// TIA Portal project "ProjektSklepu" (V18)

(* hardware
DEVICE "S7-1200 station_1"  S7-1200 Station
   slot 0: "Rack_0"  S7-1200 Rack  Rack  V1.0
   slot 1: "PLC_1"  CPU 1214C AC/DC/Rly  6ES7 214-1BG40-0XB0  V4.6
DEVICE "HMI_1"  KTP700 Basic PN
   slot 0: "HMI_1"  KTP700 Basic PN  6AV2 123-2GB03-0AX0  17.0.0.0
   slot 1: "HMI_RT_1"  KTP700 Basic PN  6AV2 123-2GB03-0AX0  17.0.0.0
   slot 5: "HMI_1.IE_CP_1"  PROFINET Interface  17.0.0.0
      slot 1: "PROFINET Interface_1"  PROFINET Interface
         slot 1: "Port_1"  Port
*)

// ===== PLC "PLC_1"  CPU 1214C AC/DC/Rly =====

VAR_GLOBAL   // PLC tag table "TT_Drzwi"
   "CzujnikRuchu_DrzwiWejscie" AT %M0.0 : Bool;
   "SygnalPracownikaDoOtwarcia_DrzwiWejscie" AT %M0.1 : Bool;
   "ZmiennaDoSymulacjiCzujnikaRuchu" AT %M0.2 : Bool;
   "StanDrzwi" AT %M0.7 : Bool;
   "Clock_Byte" AT %MB100 : Byte;
   "Clock_10Hz" AT %M100.0 : Bool;
   "Clock_5Hz" AT %M100.1 : Bool;
   "Clock_2.5Hz" AT %M100.2 : Bool;
   "Clock_2Hz" AT %M100.3 : Bool;
   "Clock_1.25Hz" AT %M100.4 : Bool;
   "Clock_1Hz" AT %M100.5 : Bool;
   "Clock_0.625Hz" AT %M100.6 : Bool;
   "Clock_0.5Hz" AT %M100.7 : Bool;
   "CzujnikRuchuWyjscie" AT %M101.0 : Bool;
   "SygnalPracownikaDoWyjscie" AT %M101.1 : Bool;
   "Liczba osob" AT %MW6 : Int;
   "zmienna pomocnicza do wentylacji" AT %M8.1 : Bool;
   "ZmiennaPomocnicza do zliczania osob" AT %M8.2 : Bool;
   "ZmiennaPomocnicza do zliczania osob wyjscie" AT %M8.3 : Bool;
   "Odliczanie" AT %M8.4 : Bool;
   "StanDrzwiINT" AT %MW4 : Int;
END_VAR

VAR_GLOBAL   // PLC tag table "TT_Temperatura"
   "Grzanie" AT %M0.3 : Bool;
   "Chłodzenie" AT %M0.4 : Bool;
   "ZmiennaPomocnicznaDoGrzania" AT %M0.5 : Bool;
   "ZmiennaPomocniczaDoChłodzenia" AT %M0.6 : Bool;
END_VAR

VAR_GLOBAL   // PLC tag table "TT_Pozar"
   "Tlo" AT %M1.0 : Bool;
   "PrzyciskDoSymulacjiCzujnikaDymu" AT %M1.1 : Bool;
   "CzujnikDymu" AT %M1.2 : Bool;
   "Swiatlo alarmowe" AT %M1.3 : Bool;
   "PracownikAlarm" AT %M1.4 : Bool;
   "ALARM" AT %M1.5 : Bool;
   "Zmienna pomocnicza do swiatla alarmu" AT %M1.6 : Bool;
   "ZmiennaDoSymulacjiCzujnikaWyjscie" AT %M1.7 : Bool;
   "Wlacz wentylacje" AT %M2.0 : Bool;
END_VAR

DATA_BLOCK "Przycisk_DB"   // DB1
{ S7_Optimized_Access := 'TRUE' }
VERSION : 0.1
// stored: InstanceOfName Przycisk
"Przycisk"
BEGIN
END_DATA_BLOCK

DATA_BLOCK "Temperatura"   // DB4
{ S7_Optimized_Access := 'TRUE' }
VERSION : 0.1
   VAR
      TemperaturaAktualna : Int := 15;
      TemperaturaDanaPrzezPracownika : Int := 15;
   END_VAR
BEGIN
END_DATA_BLOCK

DATA_BLOCK "Przycisk_DB_1"   // DB5
{ S7_Optimized_Access := 'TRUE' }
VERSION : 0.1
// stored: InstanceOfName Przycisk
"Przycisk"
BEGIN
END_DATA_BLOCK

DATA_BLOCK "Przycisk_DB_2"   // DB6
{ S7_Optimized_Access := 'TRUE' }
VERSION : 0.1
// stored: InstanceOfName Przycisk
"Przycisk"
BEGIN
END_DATA_BLOCK

DATA_BLOCK "Block_1_DB"   // DB7
{ S7_Optimized_Access := 'TRUE' }
VERSION : 0.1
// stored: InstanceOfName ZmianaBoolNaInt
"ZmianaBoolNaInt"
BEGIN
END_DATA_BLOCK

DATA_BLOCK "Przycisk_DB_3"   // DB8
{ S7_Optimized_Access := 'TRUE' }
VERSION : 0.1
// stored: InstanceOfName Przycisk
"Przycisk"
BEGIN
END_DATA_BLOCK

DATA_BLOCK "Block_1_DB_1"   // DB9
{ S7_Optimized_Access := 'TRUE' }
VERSION : 0.1
// stored: InstanceOfName ZmianaBoolNaInt
"ZmianaBoolNaInt"
BEGIN
END_DATA_BLOCK

// folder: System blocks/Program resources

DATA_BLOCK "IEC_Timer_0_DB"   // DB2
{ S7_Optimized_Access := 'TRUE' }
AUTHOR : Simatic
FAMILY : IEC
NAME : IEC_TMR
VERSION : 1.0
// stored: InstanceOfName IEC_TIMER
"IEC_TIMER"
BEGIN
END_DATA_BLOCK

DATA_BLOCK "IEC_Timer_0_DB_1"   // DB3
{ S7_Optimized_Access := 'TRUE' }
AUTHOR : Simatic
FAMILY : IEC
NAME : IEC_TMR
VERSION : 1.0
// stored: InstanceOfName IEC_TIMER
"IEC_TIMER"
BEGIN
END_DATA_BLOCK

DATA_BLOCK "IEC_Timer_0_DB_4"   // DB10
{ S7_Optimized_Access := 'TRUE' }
AUTHOR : Simatic
FAMILY : IEC
NAME : IEC_TMR
VERSION : 1.0
// stored: InstanceOfName IEC_TIMER
"IEC_TIMER"
BEGIN
END_DATA_BLOCK

// folder: (top level)

FUNCTION_BLOCK "Przycisk"   // FB1, SCL
{ S7_Optimized_Access := 'TRUE' }
VERSION : 0.1
   VAR_INPUT
      HMI_Przycisk : Bool;
   END_VAR
   VAR_IN_OUT
      Lampka : Bool;
   END_VAR
   VAR
      Prev_HMI_Button : Bool;
   END_VAR
BEGIN
   IF #HMI_Przycisk AND NOT #Prev_HMI_Button THEN
       #Lampka := NOT #Lampka;
   END_IF;

   #Prev_HMI_Button := #HMI_Przycisk;
END_FUNCTION_BLOCK

FUNCTION_BLOCK "ZmianaBoolNaInt"   // FB2, SCL
{ S7_Optimized_Access := 'TRUE' }
VERSION : 0.1
   VAR_INPUT
      StanDrzwi : Bool;
   END_VAR
   VAR_OUTPUT
      StanDrzwiInt : Int;
   END_VAR
BEGIN
   IF "StanDrzwi" THEN
       #StanDrzwiInt := 1;
   ELSE
       #StanDrzwiInt := 0;
   END_IF;
END_FUNCTION_BLOCK

ORGANIZATION_BLOCK "Main"   // OB1, LAD, ProgramCycle
TITLE = "Main Program Sweep (Cycle)"
{ S7_Optimized_Access := 'TRUE' }
VERSION : 0.1
   VAR_INPUT
      Initial_Call : Bool;   // Initial call of this OB
      Remanence : Bool;   // =True, if remanent data are available
   END_VAR
   VAR_TEMP   // added for the SCL form of the ladder/FBD networks
      _w1 : Bool;
      _w2 : Bool;
   END_VAR
BEGIN

REGION Network 1: Zmienia stan czujnika wejścia za każdym razem, gdy przycisk zostanie naciśnięty - na zbocze narastające
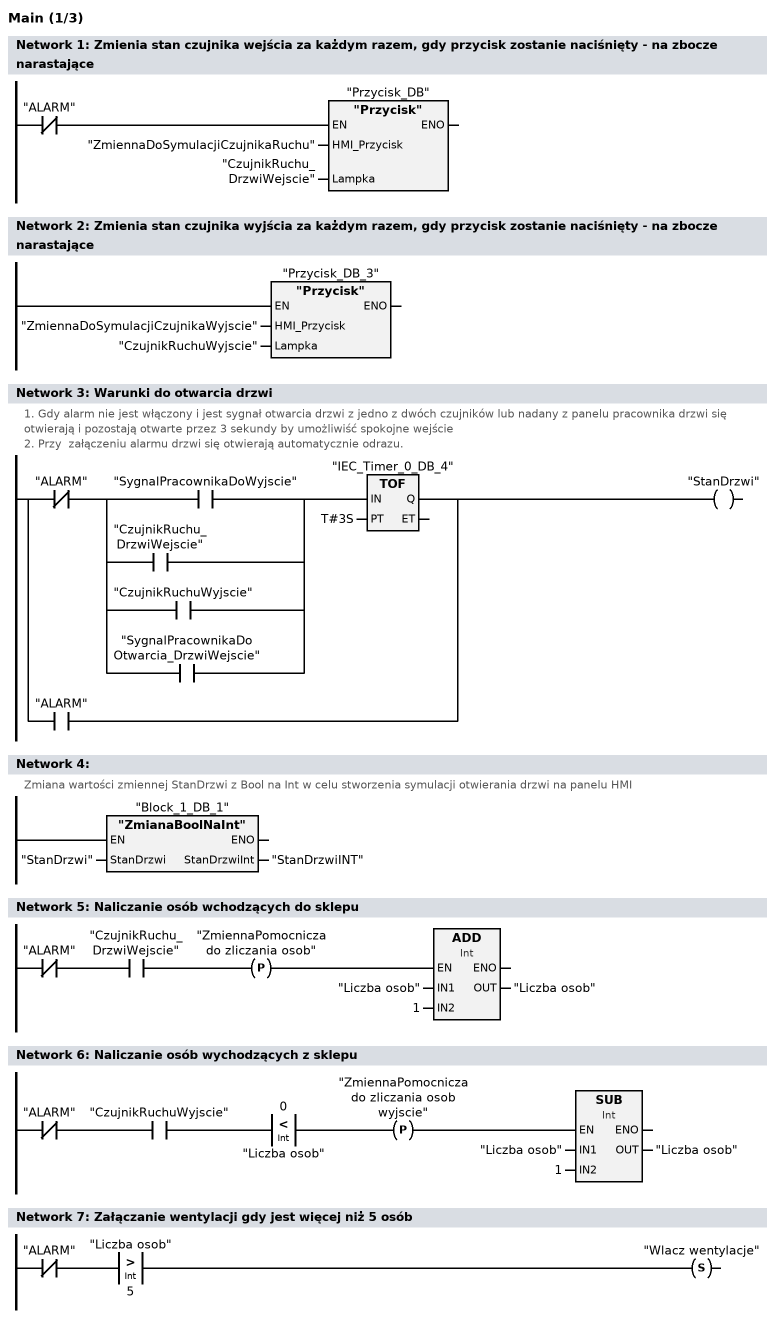
   RUNG wire#powerrail
      I_Contact( "ALARM" )
      "Przycisk_DB"(HMI_Przycisk := "ZmiennaDoSymulacjiCzujnikaRuchu", Lampka := "CzujnikRuchu_DrzwiWejscie")
   END_RUNG
   // the same network as SCL:
   IF NOT "ALARM" THEN
       "Przycisk_DB"(HMI_Przycisk := "ZmiennaDoSymulacjiCzujnikaRuchu", Lampka := "CzujnikRuchu_DrzwiWejscie");   // "Przycisk"
   END_IF;
END_REGION

REGION Network 2: Zmienia stan czujnika wyjścia za każdym razem, gdy przycisk zostanie naciśnięty - na zbocze narastające
   RUNG wire#powerrail
      "Przycisk_DB_3"(HMI_Przycisk := "ZmiennaDoSymulacjiCzujnikaWyjscie", Lampka := "CzujnikRuchuWyjscie")
   END_RUNG
   // the same network as SCL:
   "Przycisk_DB_3"(HMI_Przycisk := "ZmiennaDoSymulacjiCzujnikaWyjscie", Lampka := "CzujnikRuchuWyjscie");   // "Przycisk"
END_REGION

REGION Network 3: Warunki do otwarcia drzwi
   // 1. Gdy alarm nie jest włączony i jest sygnał otwarcia drzwi z jedno z dwóch czujników lub nadany z panelu pracownika drzwi się otwierają i pozostają otwarte przez 3 sekundy by umożliwiść spokojne wejście
   // 2. Przy  załączeniu alarmu drzwi się otwierają automatycznie odrazu.
   "IEC_Timer_0_DB_4".TOF(IN := NOT "ALARM" AND ("SygnalPracownikaDoWyjscie" OR "CzujnikRuchu_DrzwiWejscie" OR "CzujnikRuchuWyjscie" OR "SygnalPracownikaDoOtwarcia_DrzwiWejscie"),
                          PT := T#3S);
   "StanDrzwi" := "IEC_Timer_0_DB_4".Q OR "ALARM";
END_REGION

REGION Network 4
   // Zmiana wartości zmiennej StanDrzwi z Bool na Int w celu stworzenia symulacji otwierania drzwi na panelu HMI
   RUNG wire#powerrail
      "Block_1_DB_1"(StanDrzwi := "StanDrzwi", StanDrzwiInt => "StanDrzwiINT")
   END_RUNG
   // the same network as SCL:
   "Block_1_DB_1"(StanDrzwi := "StanDrzwi", StanDrzwiInt => "StanDrzwiINT");   // "ZmianaBoolNaInt"
END_REGION

REGION Network 5: Naliczanie osób wchodzących do sklepu
   RUNG wire#powerrail
      I_Contact( "ALARM" )
      Contact( "CzujnikRuchu_DrzwiWejscie" )
      P_Trig( "ZmiennaPomocnicza do zliczania osob" )
      { S7_Templates := "SrcType := Int" } Add(in1 := "Liczba osob", in2 := 1, out => "Liczba osob")
   END_RUNG
   // the same network as SCL:
   #_w1 := NOT "ALARM" AND "CzujnikRuchu_DrzwiWejscie";
   #_w2 := #_w1 AND NOT "ZmiennaPomocnicza do zliczania osob";   // rising edge
   "ZmiennaPomocnicza do zliczania osob" := #_w1;
   IF #_w2 THEN "Liczba osob" := "Liczba osob" + 1; END_IF;
END_REGION

REGION Network 6: Naliczanie osób wychodzących z sklepu
   RUNG wire#powerrail
      I_Contact( "ALARM" )
      Contact( "CzujnikRuchuWyjscie" )
      { S7_Templates := "SrcType := Int" } LT_Contact(in1 := 0, in2 := "Liczba osob")
      P_Trig( "ZmiennaPomocnicza do zliczania osob wyjscie" )
      { S7_Templates := "SrcType := Int" } Sub(in1 := "Liczba osob", in2 := 1, out => "Liczba osob")
   END_RUNG
   // the same network as SCL:
   #_w1 := NOT "ALARM" AND "CzujnikRuchuWyjscie" AND (0 < "Liczba osob");
   #_w2 := #_w1 AND NOT "ZmiennaPomocnicza do zliczania osob wyjscie";   // rising edge
   "ZmiennaPomocnicza do zliczania osob wyjscie" := #_w1;
   IF #_w2 THEN "Liczba osob" := "Liczba osob" - 1; END_IF;
END_REGION

REGION Network 7: Załączanie wentylacji gdy jest więcej niż 5 osób
   RUNG wire#powerrail
      I_Contact( "ALARM" )
      { S7_Templates := "SrcType := Int" } GT_Contact(in1 := "Liczba osob", in2 := 5)
      S_Coil( "Wlacz wentylacje" )
   END_RUNG
   // the same network as SCL:
   IF NOT "ALARM" AND ("Liczba osob" > 5) THEN "Wlacz wentylacje" := TRUE; END_IF;
END_REGION

REGION Network 8: Wyłączanie wentylacji gdy jest mniej niz 5 osób
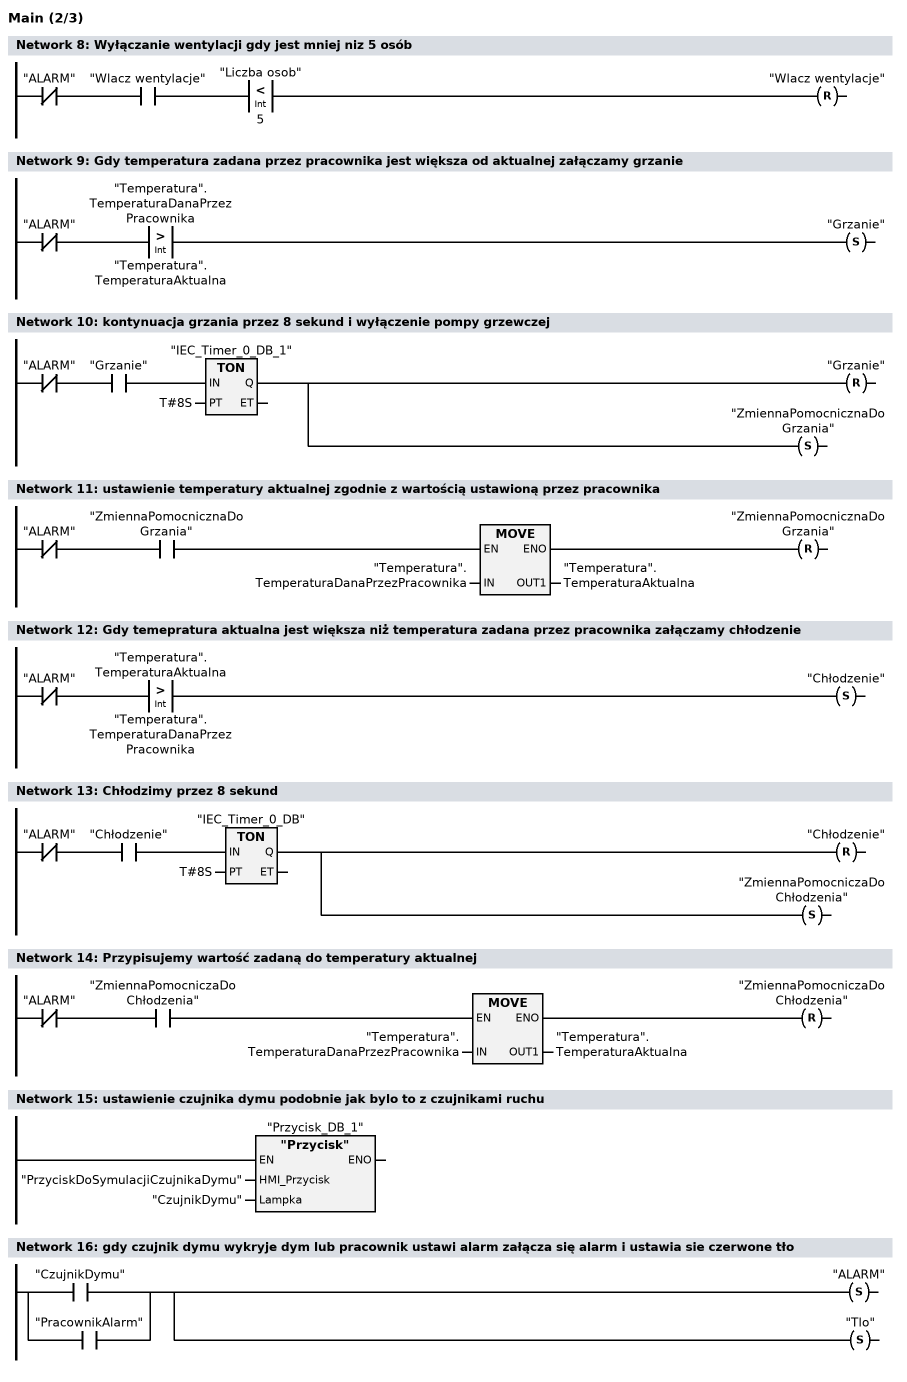
   RUNG wire#powerrail
      I_Contact( "ALARM" )
      Contact( "Wlacz wentylacje" )
      { S7_Templates := "SrcType := Int" } LT_Contact(in1 := "Liczba osob", in2 := 5)
      R_Coil( "Wlacz wentylacje" )
   END_RUNG
   // the same network as SCL:
   IF NOT "ALARM" AND "Wlacz wentylacje" AND ("Liczba osob" < 5) THEN "Wlacz wentylacje" := FALSE; END_IF;
END_REGION

REGION Network 9: Gdy temperatura zadana przez pracownika jest większa od aktualnej załączamy grzanie
   RUNG wire#powerrail
      I_Contact( "ALARM" )
      { S7_Templates := "SrcType := Int" } GT_Contact(in1 := "Temperatura".TemperaturaDanaPrzezPracownika, in2 := "Temperatura".TemperaturaAktualna)
      S_Coil( "Grzanie" )
   END_RUNG
   // the same network as SCL:
   IF NOT "ALARM" AND ("Temperatura".TemperaturaDanaPrzezPracownika > "Temperatura".TemperaturaAktualna) THEN
       "Grzanie" := TRUE;
   END_IF;
END_REGION

REGION Network 10: kontynuacja grzania przez 8 sekund i wyłączenie pompy grzewczej
   "IEC_Timer_0_DB_1".TON(IN := NOT "ALARM" AND "Grzanie", PT := T#8S);
   IF "IEC_Timer_0_DB_1".Q THEN
       "Grzanie" := FALSE;
       "ZmiennaPomocnicznaDoGrzania" := TRUE;
   END_IF;
END_REGION

REGION Network 11: ustawienie temperatury aktualnej zgodnie z wartością ustawioną przez pracownika
   RUNG wire#powerrail
      I_Contact( "ALARM" )
      Contact( "ZmiennaPomocnicznaDoGrzania" )
      Move(in := "Temperatura".TemperaturaDanaPrzezPracownika, out1 => "Temperatura".TemperaturaAktualna)
      R_Coil( "ZmiennaPomocnicznaDoGrzania" )
   END_RUNG
   // the same network as SCL:
   IF NOT "ALARM" AND "ZmiennaPomocnicznaDoGrzania" THEN
       "Temperatura".TemperaturaAktualna := "Temperatura".TemperaturaDanaPrzezPracownika;
       "ZmiennaPomocnicznaDoGrzania" := FALSE;
   END_IF;
END_REGION

REGION Network 12: Gdy temepratura aktualna jest większa niż temperatura zadana przez pracownika załączamy chłodzenie
   RUNG wire#powerrail
      I_Contact( "ALARM" )
      { S7_Templates := "SrcType := Int" } GT_Contact(in1 := "Temperatura".TemperaturaAktualna, in2 := "Temperatura".TemperaturaDanaPrzezPracownika)
      S_Coil( "Chłodzenie" )
   END_RUNG
   // the same network as SCL:
   IF NOT "ALARM" AND ("Temperatura".TemperaturaAktualna > "Temperatura".TemperaturaDanaPrzezPracownika) THEN
       "Chłodzenie" := TRUE;
   END_IF;
END_REGION

REGION Network 13: Chłodzimy przez 8 sekund
   "IEC_Timer_0_DB".TON(IN := NOT "ALARM" AND "Chłodzenie", PT := T#8S);
   IF "IEC_Timer_0_DB".Q THEN
       "Chłodzenie" := FALSE;
       "ZmiennaPomocniczaDoChłodzenia" := TRUE;
   END_IF;
END_REGION

REGION Network 14: Przypisujemy wartość zadaną do temperatury aktualnej
   RUNG wire#powerrail
      I_Contact( "ALARM" )
      Contact( "ZmiennaPomocniczaDoChłodzenia" )
      Move(in := "Temperatura".TemperaturaDanaPrzezPracownika, out1 => "Temperatura".TemperaturaAktualna)
      R_Coil( "ZmiennaPomocniczaDoChłodzenia" )
   END_RUNG
   // the same network as SCL:
   IF NOT "ALARM" AND "ZmiennaPomocniczaDoChłodzenia" THEN
       "Temperatura".TemperaturaAktualna := "Temperatura".TemperaturaDanaPrzezPracownika;
       "ZmiennaPomocniczaDoChłodzenia" := FALSE;
   END_IF;
END_REGION

REGION Network 15: ustawienie czujnika dymu podobnie jak bylo to z czujnikami ruchu
   RUNG wire#powerrail
      "Przycisk_DB_1"(HMI_Przycisk := "PrzyciskDoSymulacjiCzujnikaDymu", Lampka := "CzujnikDymu")
   END_RUNG
   // the same network as SCL:
   "Przycisk_DB_1"(HMI_Przycisk := "PrzyciskDoSymulacjiCzujnikaDymu", Lampka := "CzujnikDymu");   // "Przycisk"
END_REGION

REGION Network 16: gdy czujnik dymu wykryje dym lub pracownik ustawi alarm załącza się alarm i ustawia sie czerwone tło
   RUNG wire#powerrail
      Contact( "CzujnikDymu" )
      wire#w1
      S_Coil( "ALARM" )
   END_RUNG
   RUNG wire#powerrail
      Contact( "PracownikAlarm" )
   END_RUNG wire#w1
   RUNG wire#w1
      S_Coil( "Tlo" )
   END_RUNG
   // the same network as SCL:
   IF "CzujnikDymu" OR "PracownikAlarm" THEN
       "ALARM" := TRUE;
       "Tlo" := TRUE;
   END_IF;
END_REGION

REGION Network 17: załączamy swiatlo alarmowe ktore miga co 0.5hz zgodnie z zmienna zegarową
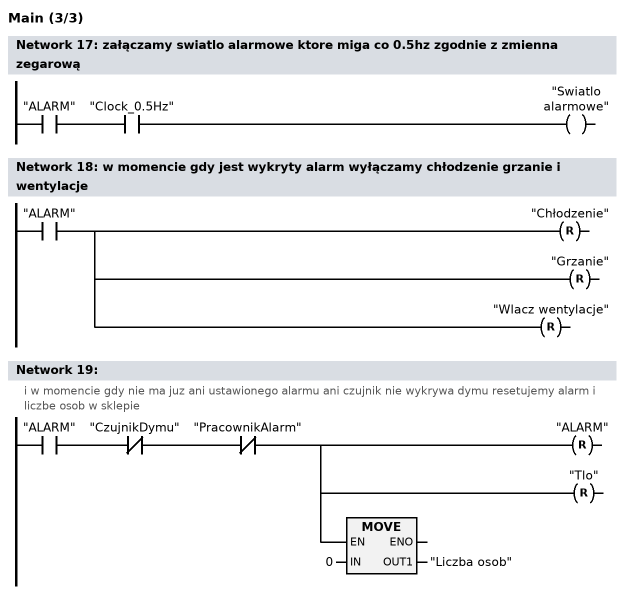
   RUNG wire#powerrail
      Contact( "ALARM" )
      Contact( "Clock_0.5Hz" )
      Coil( "Swiatlo alarmowe" )
   END_RUNG
   // the same network as SCL:
   "Swiatlo alarmowe" := "ALARM" AND "Clock_0.5Hz";
END_REGION

REGION Network 18: w momencie gdy jest wykryty alarm wyłączamy chłodzenie grzanie i wentylacje
   RUNG wire#powerrail
      Contact( "ALARM" )
      wire#w1
      R_Coil( "Chłodzenie" )
   END_RUNG
   RUNG wire#w1
      R_Coil( "Grzanie" )
   END_RUNG
   RUNG wire#w1
      R_Coil( "Wlacz wentylacje" )
   END_RUNG
   // the same network as SCL:
   IF "ALARM" THEN
       "Chłodzenie" := FALSE;
       "Grzanie" := FALSE;
       "Wlacz wentylacje" := FALSE;
   END_IF;
END_REGION

REGION Network 19
   // i w momencie gdy nie ma juz ani ustawionego alarmu ani czujnik nie wykrywa dymu resetujemy alarm i liczbe osob w sklepie
   RUNG wire#powerrail
      Contact( "ALARM" )
      I_Contact( "CzujnikDymu" )
      I_Contact( "PracownikAlarm" )
      wire#w1
      R_Coil( "ALARM" )
   END_RUNG
   RUNG wire#w1
      R_Coil( "Tlo" )
   END_RUNG
   RUNG wire#w1
      Move(in := 0, out1 => "Liczba osob")
   END_RUNG
   // the same network as SCL:
   #_w1 := "ALARM" AND NOT "CzujnikDymu" AND NOT "PracownikAlarm";
   IF #_w1 THEN
       "ALARM" := FALSE;
       "Tlo" := FALSE;
       "Liczba osob" := 0;
   END_IF;
END_REGION
END_ORGANIZATION_BLOCK

(* ===== HMI "HMI_RT_1" =====
system functions are stored by id; their names below are inferred from use
connection "HMI_Connection_1": ETHERNET, SMART_S7_1200_OMS

HMI tags "Default tag table"
   "Tag_ScreenNumber" : UInt, internal
   "ZmiennaDoSymulacjiCzujnikaRuchu" : Bool = PLC ZmiennaDoSymulacjiCzujnikaRuchu AT %M0.2, 500 ms
   "CzujnikRuchu_DrzwiWejscie" : Bool = PLC CzujnikRuchu_DrzwiWejscie AT %M0.0, 500 ms
   "SygnalPracownikaDoOtwarcia_DrzwiWejscie" : Bool = PLC SygnalPracownikaDoOtwarcia_DrzwiWejscie AT %M0.1, 500 ms
   "StanDrzwi" : Bool = PLC StanDrzwi AT %M0.7, 500 ms
   "Grzanie" : Bool = PLC Grzanie AT %M0.3, 500 ms
   "Chłodzenie" : Bool = PLC Chłodzenie AT %M0.4, 500 ms
   "Temperatura_TemperaturaAktualna" : Int = PLC Temperatura.TemperaturaAktualna, 500 ms
   "Temperatura_TemperaturaDanaPrzezPracownika" : Int = PLC Temperatura.TemperaturaDanaPrzezPracownika, 500 ms
   "PrzyciskDoSymulacjiCzujnikaDymu" : Bool = PLC PrzyciskDoSymulacjiCzujnikaDymu AT %M1.1, 500 ms
   "CzujnikDymu" : Bool = PLC CzujnikDymu AT %M1.2, 500 ms
   "PracownikAlarm" : Bool = PLC PracownikAlarm AT %M1.4, 500 ms
   "Swiatlo alarmowe" : Bool = PLC "Swiatlo alarmowe" AT %M1.3, 500 ms
   "Tlo" : Bool = PLC Tlo AT %M1.0, 500 ms
   "ZmiennaDoSymulacjiCzujnikaWyjscie" : Bool = PLC ZmiennaDoSymulacjiCzujnikaWyjscie AT %M1.7, 500 ms
   "CzujnikRuchuWyjscie" : Bool = PLC CzujnikRuchuWyjscie AT %M101.0, 500 ms
   "SygnalPracownikaDoWyjscie" : Bool = PLC SygnalPracownikaDoWyjscie AT %M101.1, 500 ms
   "Liczba osob" : Int = PLC "Liczba osob" AT %MW6, 500 ms
   "Wlacz wentylacje" : Bool = PLC "Wlacz wentylacje" AT %M2.0, 500 ms
   "StanDrzwiINT" : Int = PLC StanDrzwiINT AT %MW4, 500 ms

Template "Template_1" 800x480
   Button "Exit" at 714,429 size 71x50; TextOff 'Exit'; PictureOff "ExitRuntime_KTP700_Basic_PN_TR"; PictureOn "ExitRuntime_KTP700_Basic_PN_TR"
      on Release: StopRuntime(0)
   Button "Template_Button" at 614,429 size 71x50; TextOff 'Text'
   Button "Template_Button_1" at 514,429 size 71x50; TextOff 'Text'
   Button "Template_Button_2" at 414,429 size 71x50; TextOff 'Text'
   Button "Template_Button_3" at 314,429 size 71x50; TextOff 'Text'
   Button "Template_Button_4" at 214,429 size 71x50; TextOff 'Text'
   Button "Alarms" at 114,429 size 71x50; TextOff 'Alarms'; PictureOff "AlarmDisplay_KTP700_Basic_PN_TR"; PictureOn "AlarmDisplay_KTP700_Basic_PN_TR"
      on Release: function_ef3f5d25("Alarm window_Unacknowledged", -1)
   Button "Start screen" at 14,429 size 71x50; TextOff 'Start screen'; PictureOff "NavigateHome_KTP700_Basic_PN_TR"; PictureOn "NavigateHome_KTP700_Basic_PN_TR"
   SymbolicIOField "Symbolic_IO_Field_Screen" at 93,9 size 600x33; TextOff '0'; TextOn '1'; TextList "TextList_ScreenNames"
      ProcessValue <- "Tag_ScreenNumber"
      on Change: ActivateScreenByNumber("Tag_ScreenNumber", 0)
   DateTimeField "HmiScreenItemData" at 695,25 size 105x25
   DateTimeField "HmiScreenItemData_1" at 695,0 size 105x25
   GraphicView "Logo" at 0,0 size 91x51; Picture "Logo of HMI_1"

screen "Screen_1" 800x480
   Rectangle "Rectangle_2" at 0,0 size 799x479
      Appearance <- "Tlo"
   TextField "Text field_1" at 43,0 size 71x23; Text 'Czujniki'
   TextField "Text field_2" at 277,0 size 151x23; Text 'Panel Pracownika'
   TextField "Text field_3" at 598,0 size 161x23; Text 'Działanie urządzeń'
   Button "Button_1" at 31,38 size 88x26; TextOff 'Wejscie'
      on Press: function_b14e0dd5("ZmiennaDoSymulacjiCzujnikaRuchu", 0)
   Circle "Circle_1" at 124,36 size 33x33
      Appearance <- "CzujnikRuchu_DrzwiWejscie"
   Button "Button_2" at 261,37 size 120x24; TextOff 'Otwórz drzwi'
      on Press: SetBit("SygnalPracownikaDoOtwarcia_DrzwiWejscie")
      Appearance <- "StanDrzwi"
   Button "Button_3" at 389,37 size 124x25; TextOff 'Zamknij drzwi'
      on Press: ResetBit("SygnalPracownikaDoOtwarcia_DrzwiWejscie")
      Appearance <- "StanDrzwi"
   IOField "I/O field_1" at 329,172 size 129x46; FormatPattern 99999
      ProcessValue <- "Temperatura_TemperaturaDanaPrzezPracownika"
   TextField "Text field_4" at 288,138 size 205x23; Text 'Wprowadz temperature:'
   IOField "I/O field_2" at 42,175 size 116x40; FormatPattern s99999
      ProcessValue <- "Temperatura_TemperaturaAktualna"
   TextField "Text field_5" at 0,139 size 197x23; Text 'Aktualna Temperatura:'
   Bar "Bar_1" at 704,132 size 76x112; MinimumValue 0; MaximumValue 100
      ProcessValue <- "Temperatura_TemperaturaAktualna"
   TextField "Text field_6" at 547,152 size 79x23; Text 'Grzanie:'
   TextField "Text field_7" at 526,198 size 101x23; Text 'Chłodzenie:'
   Circle "Circle_2" at 627,143 size 39x39
      Appearance <- "Grzanie"
   Circle "Circle_3" at 627,194 size 39x39
      Appearance <- "Chłodzenie"
   Button "Button_4" at 16,303 size 117x29; TextOff 'Czujnik dymu'
      on Press: function_b14e0dd5("PrzyciskDoSymulacjiCzujnikaDymu", 0)
   Circle "Circle_4" at 146,299 size 38x38
      Appearance <- "CzujnikDymu"
   TextField "Text field_8" at 353,269 size 60x23; Text 'Alarm:'
   Circle "Circle_5" at 667,308 size 48x48
      Appearance <- "Swiatlo alarmowe"
   TextField "Text field_9" at 607,286 size 158x23; Text 'Światło alarmowe:'
   Switch "Switch_1" at 337,299 size 103x39; CaptionText 'Switch'; TextOff 'OFF'; TextOn 'ON'
      on SwitchOn: SetBit("PracownikAlarm")
      on SwitchOff: ResetBit("PracownikAlarm")
   TextField "Text field_10" at 337,388 size 96x23; Text 'Wentylacja'
   Circle "Circle_6" at 648,407 size 63x63
      Appearance <- "Wlacz wentylacje"
   Button "Button_8" at 31,77 size 88x24; TextOff 'Wyjscie'
      on Press: function_b14e0dd5("ZmiennaDoSymulacjiCzujnikaWyjscie", 0)
   Circle "Circle_7" at 125,72 size 33x33
      Appearance <- "CzujnikRuchuWyjscie"
   Button "Button_9" at 262,71 size 120x26; TextOff 'Otwórz drzwi'
      on Press: SetBit("SygnalPracownikaDoWyjscie")
      Appearance <- "StanDrzwi"
   Button "Button_10" at 389,72 size 126x26; TextOff 'Zamknij drzwi'
      on Press: ResetBit("SygnalPracownikaDoWyjscie")
      Appearance <- "StanDrzwi"
   IOField "I/O field_3" at 371,426 size 85x27; FormatPattern s99999
      ProcessValue <- "Liczba osob"
   Rectangle "Rectangle_1" at 660,38 size 30x51
      HorizontalMovement <- "StanDrzwiINT"
   Rectangle "Rectangle_3" at 687,38 size 28x51
      HorizontalMovement <- "StanDrzwiINT"
   TextField "Text field_11" at 201,427 size 158x23; Text 'Ile osob w sklepie:'
   TextField "Text field_12" at 556,54 size 58x23; Text 'Drzwi:'
   TextField "Text field_13" at 187,31 size 74x23; Text 'Wejscie:'
   TextField "Text field_14" at 190,65 size 73x23; Text 'Wyjscie:'
   TextField "Text field_15" at 625,383 size 102x23; Text 'Wentylator:'
*)